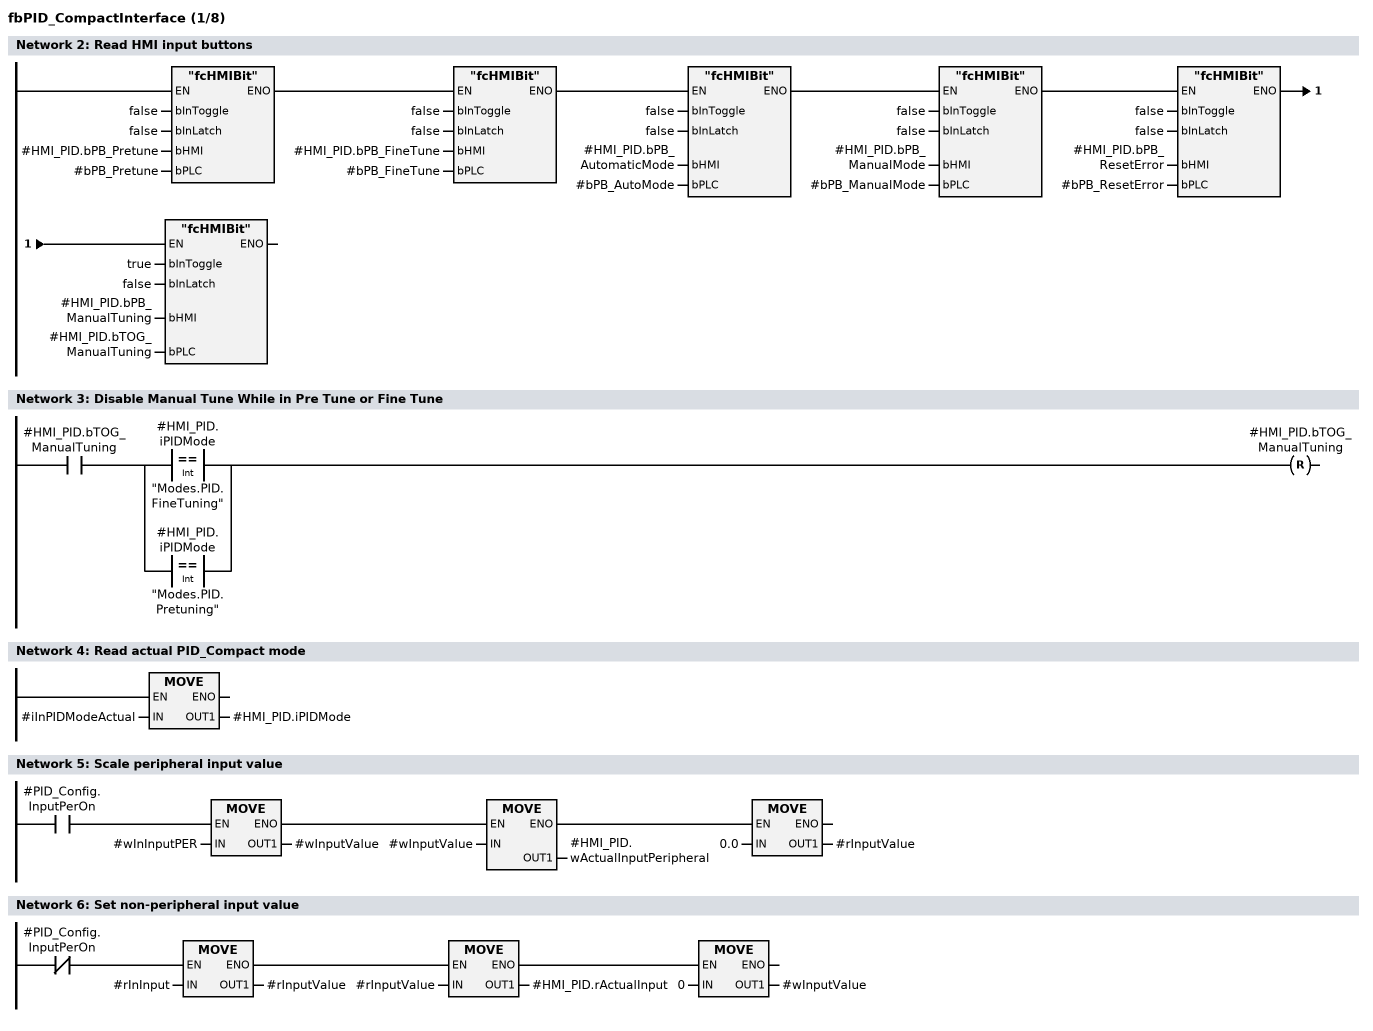
   RUNG wire#powerrail
      "fcHMIBit"(bInToggle := false, bInLatch := false, bHMI := #HMI_PID.bPB_Pretune, bPLC := #bPB_Pretune)
      "fcHMIBit"(bInToggle := false, bInLatch := false, bHMI := #HMI_PID.bPB_FineTune, bPLC := #bPB_FineTune)
      "fcHMIBit"(bInToggle := false, bInLatch := false, bHMI := #HMI_PID.bPB_AutomaticMode, bPLC := #bPB_AutoMode)
      "fcHMIBit"(bInToggle := false, bInLatch := false, bHMI := #HMI_PID.bPB_ManualMode, bPLC := #bPB_ManualMode)
      "fcHMIBit"(bInToggle := false, bInLatch := false, bHMI := #HMI_PID.bPB_ResetError, bPLC := #bPB_ResetError)
      "fcHMIBit"(bInToggle := true, bInLatch := false, bHMI := #HMI_PID.bPB_ManualTuning, bPLC := #HMI_PID.bTOG_ManualTuning)
   END_RUNG
   // the same network as SCL:
   "fcHMIBit"(bInToggle := false,
              bInLatch := false,
              bHMI := #HMI_PID.bPB_Pretune,
              bPLC := #bPB_Pretune,
              ENO => #_w1);
   "fcHMIBit"(EN := #_w1,
              bInToggle := false,
              bInLatch := false,
              bHMI := #HMI_PID.bPB_FineTune,
              bPLC := #bPB_FineTune,
              ENO => #_w2);
   "fcHMIBit"(EN := #_w2,
              bInToggle := false,
              bInLatch := false,
              bHMI := #HMI_PID.bPB_AutomaticMode,
              bPLC := #bPB_AutoMode,
              ENO => #_w3);
   "fcHMIBit"(EN := #_w3,
              bInToggle := false,
              bInLatch := false,
              bHMI := #HMI_PID.bPB_ManualMode,
              bPLC := #bPB_ManualMode,
              ENO => #_w4);
   "fcHMIBit"(EN := #_w4,
              bInToggle := false,
              bInLatch := false,
              bHMI := #HMI_PID.bPB_ResetError,
              bPLC := #bPB_ResetError,
              ENO => #_w5);
   IF #_w5 THEN
       "fcHMIBit"(bInToggle := true,
                  bInLatch := false,
                  bHMI := #HMI_PID.bPB_ManualTuning,
                  bPLC := #HMI_PID.bTOG_ManualTuning);
   END_IF;
END_REGION

REGION Network 3: Disable Manual Tune While in Pre Tune or Fine Tune
   RUNG wire#powerrail
      Contact( #HMI_PID.bTOG_ManualTuning )
      wire#w1
      { S7_Templates := "SrcType := Int" } EQ_Contact(in1 := #HMI_PID.iPIDMode, in2 := "Modes.PID.FineTuning")
      wire#w2
      R_Coil( #HMI_PID.bTOG_ManualTuning )
   END_RUNG
   RUNG wire#w1
      { S7_Templates := "SrcType := Int" } EQ_Contact(in1 := #HMI_PID.iPIDMode, in2 := "Modes.PID.Pretuning")
   END_RUNG wire#w2
   // the same network as SCL:
   IF #HMI_PID.bTOG_ManualTuning AND ((#HMI_PID.iPIDMode = "Modes.PID.FineTuning") OR (#HMI_PID.iPIDMode = "Modes.PID.Pretuning")) THEN
       #HMI_PID.bTOG_ManualTuning := FALSE;
   END_IF;
END_REGION

REGION Network 4: Read actual PID_Compact mode
   RUNG wire#powerrail
      Move(in := #iInPIDModeActual, out1 => #HMI_PID.iPIDMode)
   END_RUNG
   // the same network as SCL:
   #HMI_PID.iPIDMode := #iInPIDModeActual;
END_REGION

REGION Network 5: Scale peripheral input value
   RUNG wire#powerrail
      Contact( #PID_Config.InputPerOn )
      Move(in := #wInInputPER, out1 => #wInputValue)
      Move(in := #wInputValue, out1 => #HMI_PID.wActualInputPeripheral)
      Move(in := 0.0, out1 => #rInputValue)
   END_RUNG
   // the same network as SCL:
   IF #PID_Config.InputPerOn THEN
       #wInputValue := #wInInputPER;
       #HMI_PID.wActualInputPeripheral := #wInputValue;
       #rInputValue := 0.0;
   END_IF;
END_REGION

REGION Network 6: Set non-peripheral input value
   RUNG wire#powerrail
      I_Contact( #PID_Config.InputPerOn )
      Move(in := #rInInput, out1 => #rInputValue)
      Move(in := #rInputValue, out1 => #HMI_PID.rActualInput)
      Move(in := 0, out1 => #wInputValue)
   END_RUNG
   // the same network as SCL:
   IF NOT #PID_Config.InputPerOn THEN
       #rInputValue := #rInInput;
       #HMI_PID.rActualInput := #rInputValue;
       #wInputValue := 0;
   END_IF;
END_REGION

REGION Network 7: Check HMI tuning parameters for changes
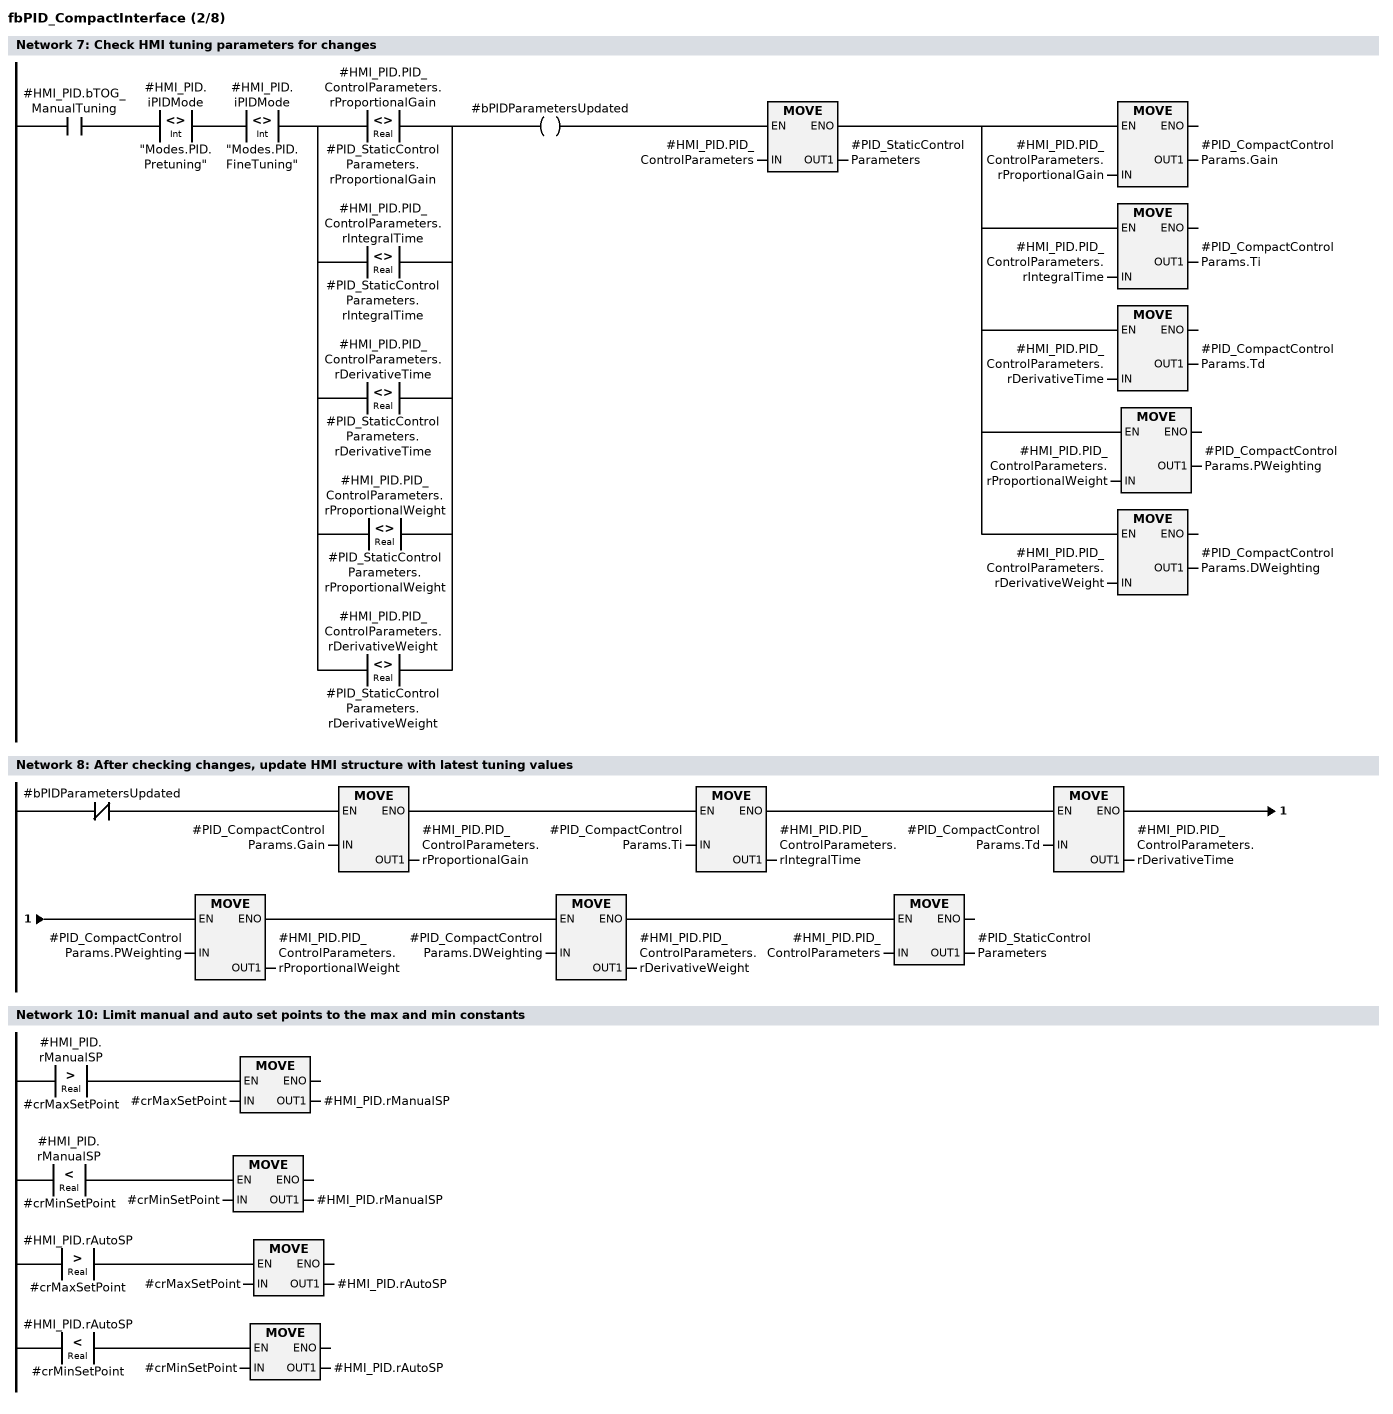
   RUNG wire#powerrail
      Contact( #HMI_PID.bTOG_ManualTuning )
      { S7_Templates := "SrcType := Int" } NE_Contact(in1 := #HMI_PID.iPIDMode, in2 := "Modes.PID.Pretuning")
      { S7_Templates := "SrcType := Int" } NE_Contact(in1 := #HMI_PID.iPIDMode, in2 := "Modes.PID.FineTuning")
      wire#w1
      { S7_Templates := "SrcType := Real" } NE_Contact(in1 := #HMI_PID.PID_ControlParameters.rProportionalGain, in2 := #PID_StaticControlParameters.rProportionalGain)
      wire#w2
      Coil( #bPIDParametersUpdated )
      Move(in := #HMI_PID.PID_ControlParameters, out1 => #PID_StaticControlParameters)
      wire#w3
      Move(in := #HMI_PID.PID_ControlParameters.rProportionalGain, out1 => #PID_CompactControlParams.Gain)
   END_RUNG
   RUNG wire#w1
      { S7_Templates := "SrcType := Real" } NE_Contact(in1 := #HMI_PID.PID_ControlParameters.rIntegralTime, in2 := #PID_StaticControlParameters.rIntegralTime)
   END_RUNG wire#w2
   RUNG wire#w1
      { S7_Templates := "SrcType := Real" } NE_Contact(in1 := #HMI_PID.PID_ControlParameters.rDerivativeTime, in2 := #PID_StaticControlParameters.rDerivativeTime)
   END_RUNG wire#w2
   RUNG wire#w1
      { S7_Templates := "SrcType := Real" } NE_Contact(in1 := #HMI_PID.PID_ControlParameters.rProportionalWeight, in2 := #PID_StaticControlParameters.rProportionalWeight)
   END_RUNG wire#w2
   RUNG wire#w1
      { S7_Templates := "SrcType := Real" } NE_Contact(in1 := #HMI_PID.PID_ControlParameters.rDerivativeWeight, in2 := #PID_StaticControlParameters.rDerivativeWeight)
   END_RUNG wire#w2
   RUNG wire#w3
      Move(in := #HMI_PID.PID_ControlParameters.rIntegralTime, out1 => #PID_CompactControlParams.Ti)
   END_RUNG
   RUNG wire#w3
      Move(in := #HMI_PID.PID_ControlParameters.rDerivativeTime, out1 => #PID_CompactControlParams.Td)
   END_RUNG
   RUNG wire#w3
      Move(in := #HMI_PID.PID_ControlParameters.rProportionalWeight, out1 => #PID_CompactControlParams.PWeighting)
   END_RUNG
   RUNG wire#w3
      Move(in := #HMI_PID.PID_ControlParameters.rDerivativeWeight, out1 => #PID_CompactControlParams.DWeighting)
   END_RUNG
   // the same network as SCL:
   #bPIDParametersUpdated := #HMI_PID.bTOG_ManualTuning AND (#HMI_PID.iPIDMode <> "Modes.PID.Pretuning") AND (#HMI_PID.iPIDMode <> "Modes.PID.FineTuning") AND ((#HMI_PID.PID_ControlParameters.rProportionalGain <> #PID_StaticControlParameters.rProportionalGain) OR (#HMI_PID.PID_ControlParameters.rIntegralTime <> #PID_StaticControlParameters.rIntegralTime) OR (#HMI_PID.PID_ControlParameters.rDerivativeTime <> #PID_StaticControlParameters.rDerivativeTime) OR (#HMI_PID.PID_ControlParameters.rProportionalWeight <> #PID_StaticControlParameters.rProportionalWeight) OR (#HMI_PID.PID_ControlParameters.rDerivativeWeight <> #PID_StaticControlParameters.rDerivativeWeight));
   IF #bPIDParametersUpdated THEN
       #PID_StaticControlParameters := #HMI_PID.PID_ControlParameters;
       #PID_CompactControlParams.Gain := #HMI_PID.PID_ControlParameters.rProportionalGain;
       #PID_CompactControlParams.Ti := #HMI_PID.PID_ControlParameters.rIntegralTime;
       #PID_CompactControlParams.Td := #HMI_PID.PID_ControlParameters.rDerivativeTime;
       #PID_CompactControlParams.PWeighting := #HMI_PID.PID_ControlParameters.rProportionalWeight;
       #PID_CompactControlParams.DWeighting := #HMI_PID.PID_ControlParameters.rDerivativeWeight;
   END_IF;
END_REGION

REGION Network 8: After checking changes, update HMI structure with latest tuning values
   RUNG wire#powerrail
      I_Contact( #bPIDParametersUpdated )
      Move(in := #PID_CompactControlParams.Gain, out1 => #HMI_PID.PID_ControlParameters.rProportionalGain)
      Move(in := #PID_CompactControlParams.Ti, out1 => #HMI_PID.PID_ControlParameters.rIntegralTime)
      Move(in := #PID_CompactControlParams.Td, out1 => #HMI_PID.PID_ControlParameters.rDerivativeTime)
      Move(in := #PID_CompactControlParams.PWeighting, out1 => #HMI_PID.PID_ControlParameters.rProportionalWeight)
      Move(in := #PID_CompactControlParams.DWeighting, out1 => #HMI_PID.PID_ControlParameters.rDerivativeWeight)
      Move(in := #HMI_PID.PID_ControlParameters, out1 => #PID_StaticControlParameters)
   END_RUNG
   // the same network as SCL:
   IF NOT #bPIDParametersUpdated THEN
       #HMI_PID.PID_ControlParameters.rProportionalGain := #PID_CompactControlParams.Gain;
       #HMI_PID.PID_ControlParameters.rIntegralTime := #PID_CompactControlParams.Ti;
       #HMI_PID.PID_ControlParameters.rDerivativeTime := #PID_CompactControlParams.Td;
       #HMI_PID.PID_ControlParameters.rProportionalWeight := #PID_CompactControlParams.PWeighting;
       #HMI_PID.PID_ControlParameters.rDerivativeWeight := #PID_CompactControlParams.DWeighting;
       #PID_StaticControlParameters := #HMI_PID.PID_ControlParameters;
   END_IF;
END_REGION

REGION Network 9: --------------------------------------------------- Control Logic ------------------------------------------------------------
END_REGION

REGION Network 10: Limit manual and auto set points to the max and min constants
   RUNG wire#powerrail
      { S7_Templates := "SrcType := Real" } GT_Contact(in1 := #HMI_PID.rManualSP, in2 := #crMaxSetPoint)
      { S7_GenerateENO := "TRUE" } Move(in := #crMaxSetPoint, out1 => #HMI_PID.rManualSP)
   END_RUNG
   RUNG wire#powerrail
      { S7_Templates := "SrcType := Real" } LT_Contact(in1 := #HMI_PID.rManualSP, in2 := #crMinSetPoint)
      { S7_GenerateENO := "TRUE" } Move(in := #crMinSetPoint, out1 => #HMI_PID.rManualSP)
   END_RUNG
   RUNG wire#powerrail
      { S7_Templates := "SrcType := Real" } GT_Contact(in1 := #HMI_PID.rAutoSP, in2 := #crMaxSetPoint)
      { S7_GenerateENO := "TRUE" } Move(in := #crMaxSetPoint, out1 => #HMI_PID.rAutoSP)
   END_RUNG
   RUNG wire#powerrail
      { S7_Templates := "SrcType := Real" } LT_Contact(in1 := #HMI_PID.rAutoSP, in2 := #crMinSetPoint)
      { S7_GenerateENO := "TRUE" } Move(in := #crMinSetPoint, out1 => #HMI_PID.rAutoSP)
   END_RUNG
   // the same network as SCL:
   IF #HMI_PID.rManualSP > #crMaxSetPoint THEN #HMI_PID.rManualSP := #crMaxSetPoint; END_IF;
   IF #HMI_PID.rManualSP < #crMinSetPoint THEN #HMI_PID.rManualSP := #crMinSetPoint; END_IF;
   IF #HMI_PID.rAutoSP > #crMaxSetPoint THEN #HMI_PID.rAutoSP := #crMaxSetPoint; END_IF;
   IF #HMI_PID.rAutoSP < #crMinSetPoint THEN #HMI_PID.rAutoSP := #crMinSetPoint; END_IF;
END_REGION

REGION Network 11: Reset errors
   // Clear all errors
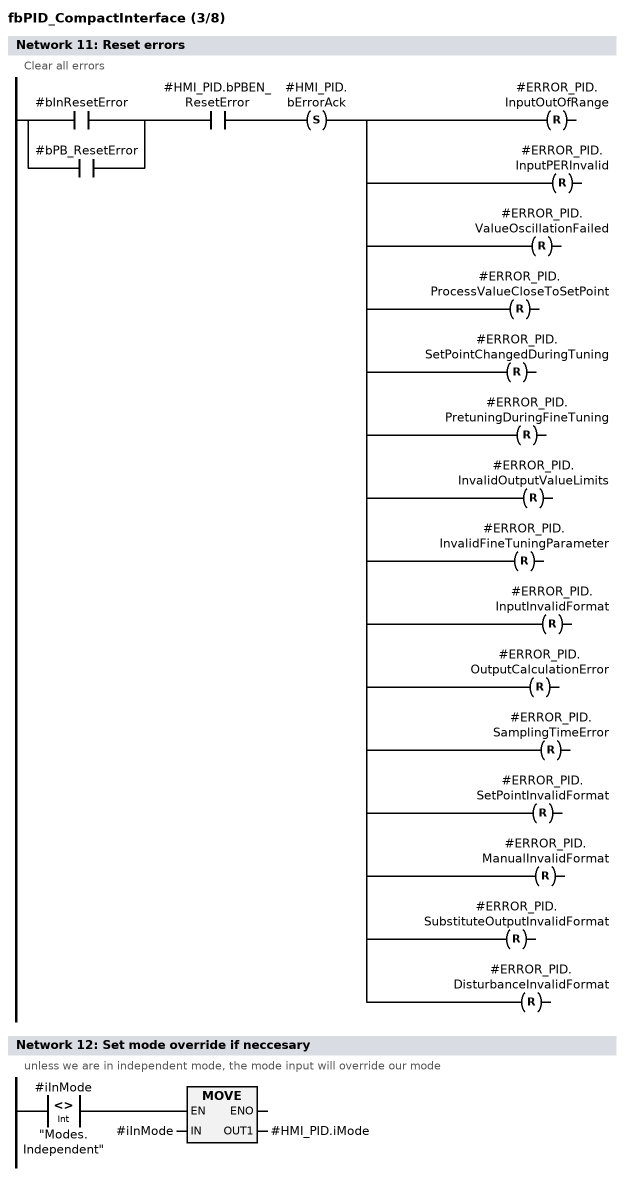
   RUNG wire#powerrail
      Contact( #bInResetError )
      wire#w1
      Contact( #HMI_PID.bPBEN_ResetError )
      S_Coil( #HMI_PID.bErrorAck )
      wire#w2
      R_Coil( #ERROR_PID.InputOutOfRange )
   END_RUNG
   RUNG wire#powerrail
      Contact( #bPB_ResetError )
   END_RUNG wire#w1
   RUNG wire#w2
      R_Coil( #ERROR_PID.InputPERInvalid )
   END_RUNG
   RUNG wire#w2
      R_Coil( #ERROR_PID.ValueOscillationFailed )
   END_RUNG
   RUNG wire#w2
      R_Coil( #ERROR_PID.ProcessValueCloseToSetPoint )
   END_RUNG
   RUNG wire#w2
      R_Coil( #ERROR_PID.SetPointChangedDuringTuning )
   END_RUNG
   RUNG wire#w2
      R_Coil( #ERROR_PID.PretuningDuringFineTuning )
   END_RUNG
   RUNG wire#w2
      R_Coil( #ERROR_PID.InvalidOutputValueLimits )
   END_RUNG
   RUNG wire#w2
      R_Coil( #ERROR_PID.InvalidFineTuningParameter )
   END_RUNG
   RUNG wire#w2
      R_Coil( #ERROR_PID.InputInvalidFormat )
   END_RUNG
   RUNG wire#w2
      R_Coil( #ERROR_PID.OutputCalculationError )
   END_RUNG
   RUNG wire#w2
      R_Coil( #ERROR_PID.SamplingTimeError )
   END_RUNG
   RUNG wire#w2
      R_Coil( #ERROR_PID.SetPointInvalidFormat )
   END_RUNG
   RUNG wire#w2
      R_Coil( #ERROR_PID.ManualInvalidFormat )
   END_RUNG
   RUNG wire#w2
      R_Coil( #ERROR_PID.SubstituteOutputInvalidFormat )
   END_RUNG
   RUNG wire#w2
      R_Coil( #ERROR_PID.DisturbanceInvalidFormat )
   END_RUNG
   // the same network as SCL:
   IF (#bInResetError OR #bPB_ResetError) AND #HMI_PID.bPBEN_ResetError THEN
       #HMI_PID.bErrorAck := TRUE;
       #ERROR_PID.InputOutOfRange := FALSE;
       #ERROR_PID.InputPERInvalid := FALSE;
       #ERROR_PID.ValueOscillationFailed := FALSE;
       #ERROR_PID.ProcessValueCloseToSetPoint := FALSE;
       #ERROR_PID.SetPointChangedDuringTuning := FALSE;
       #ERROR_PID.PretuningDuringFineTuning := FALSE;
       #ERROR_PID.InvalidOutputValueLimits := FALSE;
       #ERROR_PID.InvalidFineTuningParameter := FALSE;
       #ERROR_PID.InputInvalidFormat := FALSE;
       #ERROR_PID.OutputCalculationError := FALSE;
       #ERROR_PID.SamplingTimeError := FALSE;
       #ERROR_PID.SetPointInvalidFormat := FALSE;
       #ERROR_PID.ManualInvalidFormat := FALSE;
       #ERROR_PID.SubstituteOutputInvalidFormat := FALSE;
       #ERROR_PID.DisturbanceInvalidFormat := FALSE;
   END_IF;
END_REGION

REGION Network 12: Set mode override if neccesary
   // unless we are in independent mode, the mode input will override our mode
   RUNG wire#powerrail
      { S7_Templates := "SrcType := Int" } NE_Contact(in1 := #iInMode, in2 := "Modes.Independent")
      { S7_GenerateENO := "TRUE" } Move(in := #iInMode, out1 => #HMI_PID.iMode)
   END_RUNG
   // the same network as SCL:
   IF #iInMode <> "Modes.Independent" THEN #HMI_PID.iMode := #iInMode; END_IF;
END_REGION

REGION Network 13: Determine if auto or manual mode is active
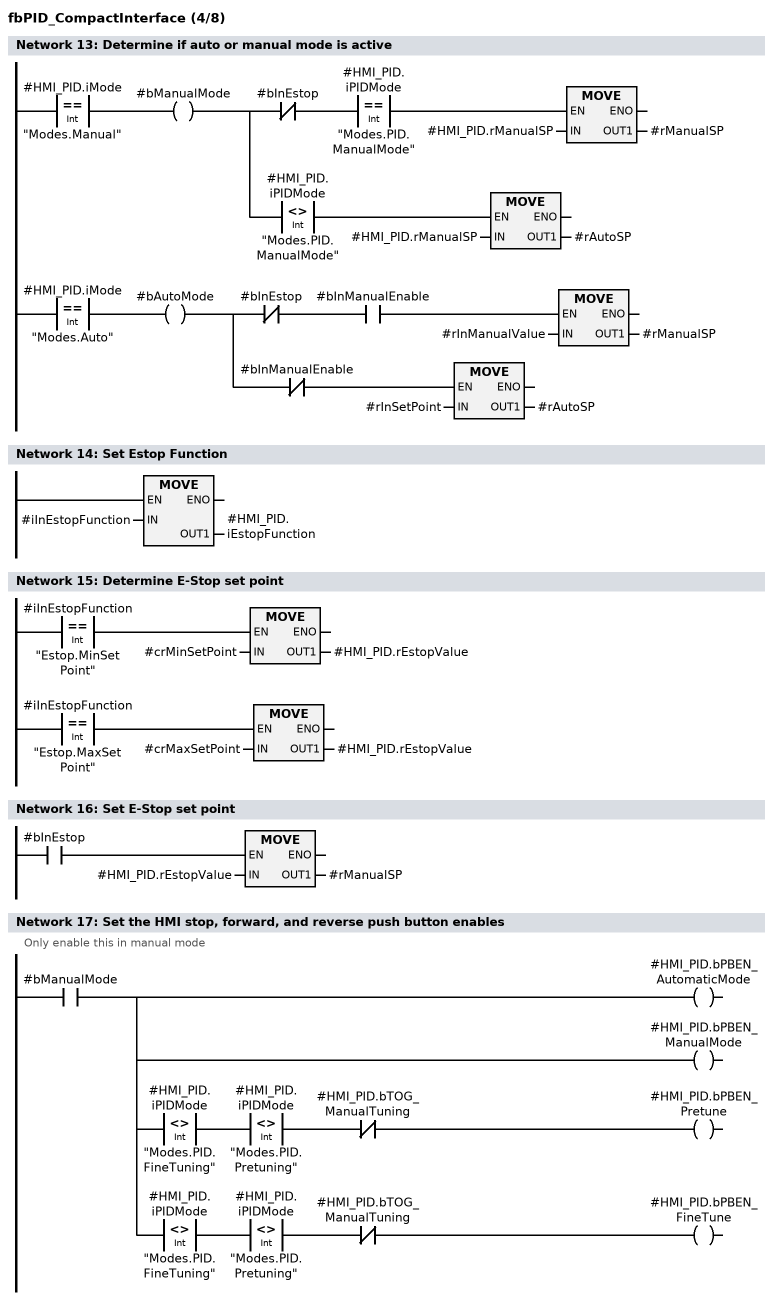
   RUNG wire#powerrail
      { S7_Templates := "SrcType := Int" } EQ_Contact(in1 := #HMI_PID.iMode, in2 := "Modes.Manual")
      Coil( #bManualMode )
      wire#w1
      I_Contact( #bInEstop )
      { S7_Templates := "SrcType := Int" } EQ_Contact(in1 := #HMI_PID.iPIDMode, in2 := "Modes.PID.ManualMode")
      { S7_GenerateENO := "TRUE" } Move(in := #HMI_PID.rManualSP, out1 => #rManualSP)
   END_RUNG
   RUNG wire#w1
      { S7_Templates := "SrcType := Int" } NE_Contact(in1 := #HMI_PID.iPIDMode, in2 := "Modes.PID.ManualMode")
      { S7_GenerateENO := "TRUE" } Move(in := #HMI_PID.rManualSP, out1 => #rAutoSP)
   END_RUNG
   RUNG wire#powerrail
      { S7_Templates := "SrcType := Int" } EQ_Contact(in1 := #HMI_PID.iMode, in2 := "Modes.Auto")
      Coil( #bAutoMode )
      wire#w2
      I_Contact( #bInEstop )
      Contact( #bInManualEnable )
      { S7_GenerateENO := "TRUE" } Move(in := #rInManualValue, out1 => #rManualSP)
   END_RUNG
   RUNG wire#w2
      I_Contact( #bInManualEnable )
      { S7_GenerateENO := "TRUE" } Move(in := #rInSetPoint, out1 => #rAutoSP)
   END_RUNG
   // the same network as SCL:
   #bManualMode := #HMI_PID.iMode = "Modes.Manual";
   IF #bManualMode AND NOT #bInEstop AND (#HMI_PID.iPIDMode = "Modes.PID.ManualMode") THEN
       #rManualSP := #HMI_PID.rManualSP;
   END_IF;
   IF #bManualMode AND (#HMI_PID.iPIDMode <> "Modes.PID.ManualMode") THEN
       #rAutoSP := #HMI_PID.rManualSP;
   END_IF;
   #bAutoMode := #HMI_PID.iMode = "Modes.Auto";
   IF #bAutoMode AND NOT #bInEstop AND #bInManualEnable THEN #rManualSP := #rInManualValue; END_IF;
   IF #bAutoMode AND NOT #bInManualEnable THEN #rAutoSP := #rInSetPoint; END_IF;
END_REGION

REGION Network 14: Set Estop Function
   RUNG wire#powerrail
      Move(in := #iInEstopFunction, out1 => #HMI_PID.iEstopFunction)
   END_RUNG
   // the same network as SCL:
   #HMI_PID.iEstopFunction := #iInEstopFunction;
END_REGION

REGION Network 15: Determine E-Stop set point
   RUNG wire#powerrail
      { S7_Templates := "SrcType := Int" } EQ_Contact(in1 := #iInEstopFunction, in2 := "Estop.MinSetPoint")
      { S7_GenerateENO := "TRUE" } Move(in := #crMinSetPoint, out1 => #HMI_PID.rEstopValue)
   END_RUNG
   RUNG wire#powerrail
      { S7_Templates := "SrcType := Int" } EQ_Contact(in1 := #iInEstopFunction, in2 := "Estop.MaxSetPoint")
      { S7_GenerateENO := "TRUE" } Move(in := #crMaxSetPoint, out1 => #HMI_PID.rEstopValue)
   END_RUNG
   // the same network as SCL:
   IF #iInEstopFunction = "Estop.MinSetPoint" THEN #HMI_PID.rEstopValue := #crMinSetPoint; END_IF;
   IF #iInEstopFunction = "Estop.MaxSetPoint" THEN #HMI_PID.rEstopValue := #crMaxSetPoint; END_IF;
END_REGION

REGION Network 16: Set E-Stop set point
   RUNG wire#powerrail
      Contact( #bInEstop )
      { S7_GenerateENO := "TRUE" } Move(in := #HMI_PID.rEstopValue, out1 => #rManualSP)
   END_RUNG
   // the same network as SCL:
   IF #bInEstop THEN #rManualSP := #HMI_PID.rEstopValue; END_IF;
END_REGION

REGION Network 17: Set the HMI stop, forward, and reverse push button enables
   // Only enable this in manual mode
   RUNG wire#powerrail
      Contact( #bManualMode )
      wire#w1
      Coil( #HMI_PID.bPBEN_AutomaticMode )
   END_RUNG
   RUNG wire#w1
      Coil( #HMI_PID.bPBEN_ManualMode )
   END_RUNG
   RUNG wire#w1
      { S7_Templates := "SrcType := Int" } NE_Contact(in1 := #HMI_PID.iPIDMode, in2 := "Modes.PID.FineTuning")
      { S7_Templates := "SrcType := Int" } NE_Contact(in1 := #HMI_PID.iPIDMode, in2 := "Modes.PID.Pretuning")
      I_Contact( #HMI_PID.bTOG_ManualTuning )
      Coil( #HMI_PID.bPBEN_Pretune )
   END_RUNG
   RUNG wire#w1
      { S7_Templates := "SrcType := Int" } NE_Contact(in1 := #HMI_PID.iPIDMode, in2 := "Modes.PID.FineTuning")
      { S7_Templates := "SrcType := Int" } NE_Contact(in1 := #HMI_PID.iPIDMode, in2 := "Modes.PID.Pretuning")
      I_Contact( #HMI_PID.bTOG_ManualTuning )
      Coil( #HMI_PID.bPBEN_FineTune )
   END_RUNG
   // the same network as SCL:
   #HMI_PID.bPBEN_AutomaticMode := #bManualMode;
   #HMI_PID.bPBEN_ManualMode := #bManualMode;
   #HMI_PID.bPBEN_Pretune := #bManualMode AND (#HMI_PID.iPIDMode <> "Modes.PID.FineTuning") AND (#HMI_PID.iPIDMode <> "Modes.PID.Pretuning") AND NOT #HMI_PID.bTOG_ManualTuning;
   #HMI_PID.bPBEN_FineTune := #bManualMode AND (#HMI_PID.iPIDMode <> "Modes.PID.FineTuning") AND (#HMI_PID.iPIDMode <> "Modes.PID.Pretuning") AND NOT #HMI_PID.bTOG_ManualTuning;
END_REGION

REGION Network 18: Enable the reset error pushbutton if there is an error
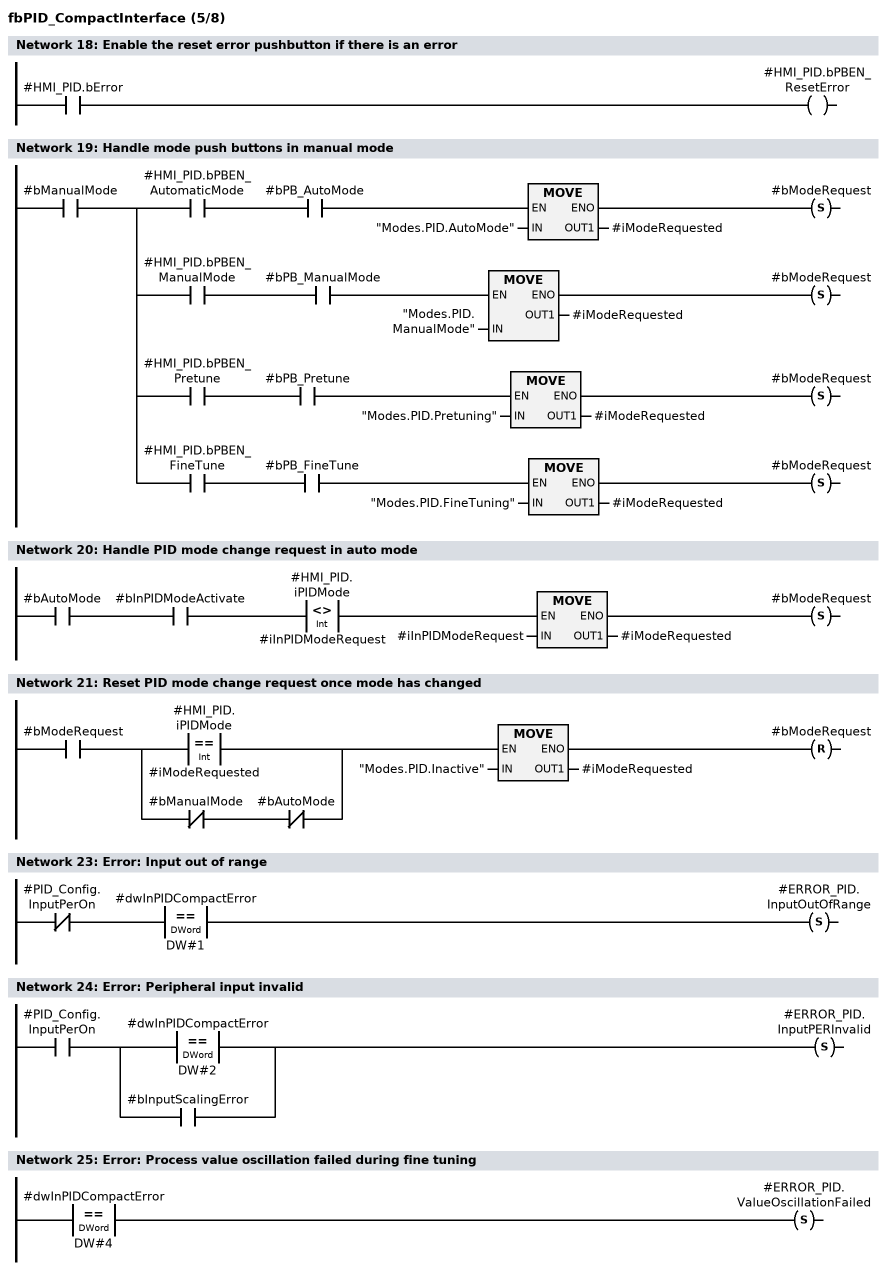
   RUNG wire#powerrail
      Contact( #HMI_PID.bError )
      Coil( #HMI_PID.bPBEN_ResetError )
   END_RUNG
   // the same network as SCL:
   #HMI_PID.bPBEN_ResetError := #HMI_PID.bError;
END_REGION

REGION Network 19: Handle mode push buttons in manual mode
   RUNG wire#powerrail
      Contact( #bManualMode )
      wire#w1
      Contact( #HMI_PID.bPBEN_AutomaticMode )
      Contact( #bPB_AutoMode )
      Move(in := "Modes.PID.AutoMode", out1 => #iModeRequested)
      S_Coil( #bModeRequest )
   END_RUNG
   RUNG wire#w1
      Contact( #HMI_PID.bPBEN_ManualMode )
      Contact( #bPB_ManualMode )
      Move(in := "Modes.PID.ManualMode", out1 => #iModeRequested)
      S_Coil( #bModeRequest )
   END_RUNG
   RUNG wire#w1
      Contact( #HMI_PID.bPBEN_Pretune )
      Contact( #bPB_Pretune )
      Move(in := "Modes.PID.Pretuning", out1 => #iModeRequested)
      S_Coil( #bModeRequest )
   END_RUNG
   RUNG wire#w1
      Contact( #HMI_PID.bPBEN_FineTune )
      Contact( #bPB_FineTune )
      Move(in := "Modes.PID.FineTuning", out1 => #iModeRequested)
      S_Coil( #bModeRequest )
   END_RUNG
   // the same network as SCL:
   IF #bManualMode AND #HMI_PID.bPBEN_AutomaticMode AND #bPB_AutoMode THEN
       #iModeRequested := "Modes.PID.AutoMode";
       #bModeRequest := TRUE;
   END_IF;
   IF #bManualMode AND #HMI_PID.bPBEN_ManualMode AND #bPB_ManualMode THEN
       #iModeRequested := "Modes.PID.ManualMode";
       #bModeRequest := TRUE;
   END_IF;
   IF #bManualMode AND #HMI_PID.bPBEN_Pretune AND #bPB_Pretune THEN
       #iModeRequested := "Modes.PID.Pretuning";
       #bModeRequest := TRUE;
   END_IF;
   IF #bManualMode AND #HMI_PID.bPBEN_FineTune AND #bPB_FineTune THEN
       #iModeRequested := "Modes.PID.FineTuning";
       #bModeRequest := TRUE;
   END_IF;
END_REGION

REGION Network 20: Handle PID mode change request in auto mode
   RUNG wire#powerrail
      Contact( #bAutoMode )
      Contact( #bInPIDModeActivate )
      { S7_Templates := "SrcType := Int" } NE_Contact(in1 := #HMI_PID.iPIDMode, in2 := #iInPIDModeRequest)
      Move(in := #iInPIDModeRequest, out1 => #iModeRequested)
      S_Coil( #bModeRequest )
   END_RUNG
   // the same network as SCL:
   IF #bAutoMode AND #bInPIDModeActivate AND (#HMI_PID.iPIDMode <> #iInPIDModeRequest) THEN
       #iModeRequested := #iInPIDModeRequest;
       #bModeRequest := TRUE;
   END_IF;
END_REGION

REGION Network 21: Reset PID mode change request once mode has changed
   RUNG wire#powerrail
      Contact( #bModeRequest )
      wire#w1
      { S7_Templates := "SrcType := Int" } EQ_Contact(in1 := #HMI_PID.iPIDMode, in2 := #iModeRequested)
      wire#w2
      Move(in := "Modes.PID.Inactive", out1 => #iModeRequested)
      R_Coil( #bModeRequest )
   END_RUNG
   RUNG wire#w1
      I_Contact( #bManualMode )
      I_Contact( #bAutoMode )
   END_RUNG wire#w2
   // the same network as SCL:
   #_w1 := #bModeRequest AND ((#HMI_PID.iPIDMode = #iModeRequested) OR (NOT #bManualMode AND NOT #bAutoMode));
   IF #_w1 THEN
       #iModeRequested := "Modes.PID.Inactive";
       #bModeRequest := FALSE;
   END_IF;
END_REGION

REGION Network 22: --------------------------------------------------------- Errors ------------------------------------------------------------------
END_REGION

REGION Network 23: Error: Input out of range
   RUNG wire#powerrail
      I_Contact( #PID_Config.InputPerOn )
      { S7_Templates := "SrcType := DWord" } EQ_Contact(in1 := #dwInPIDCompactError, in2 := DW#1)
      S_Coil( #ERROR_PID.InputOutOfRange )
   END_RUNG
   // the same network as SCL:
   IF NOT #PID_Config.InputPerOn AND (#dwInPIDCompactError = DW#1) THEN
       #ERROR_PID.InputOutOfRange := TRUE;
   END_IF;
END_REGION

REGION Network 24: Error: Peripheral input invalid
   RUNG wire#powerrail
      Contact( #PID_Config.InputPerOn )
      wire#w1
      { S7_Templates := "SrcType := DWord" } EQ_Contact(in1 := #dwInPIDCompactError, in2 := DW#2)
      wire#w2
      S_Coil( #ERROR_PID.InputPERInvalid )
   END_RUNG
   RUNG wire#w1
      Contact( #bInputScalingError )
   END_RUNG wire#w2
   // the same network as SCL:
   IF #PID_Config.InputPerOn AND ((#dwInPIDCompactError = DW#2) OR #bInputScalingError) THEN
       #ERROR_PID.InputPERInvalid := TRUE;
   END_IF;
END_REGION

REGION Network 25: Error: Process value oscillation failed during fine tuning
   RUNG wire#powerrail
      { S7_Templates := "SrcType := DWord" } EQ_Contact(in1 := #dwInPIDCompactError, in2 := DW#4)
      S_Coil( #ERROR_PID.ValueOscillationFailed )
   END_RUNG
   // the same network as SCL:
   IF #dwInPIDCompactError = DW#4 THEN #ERROR_PID.ValueOscillationFailed := TRUE; END_IF;
END_REGION

REGION Network 26: Error: Process value too close to set point for pretuning
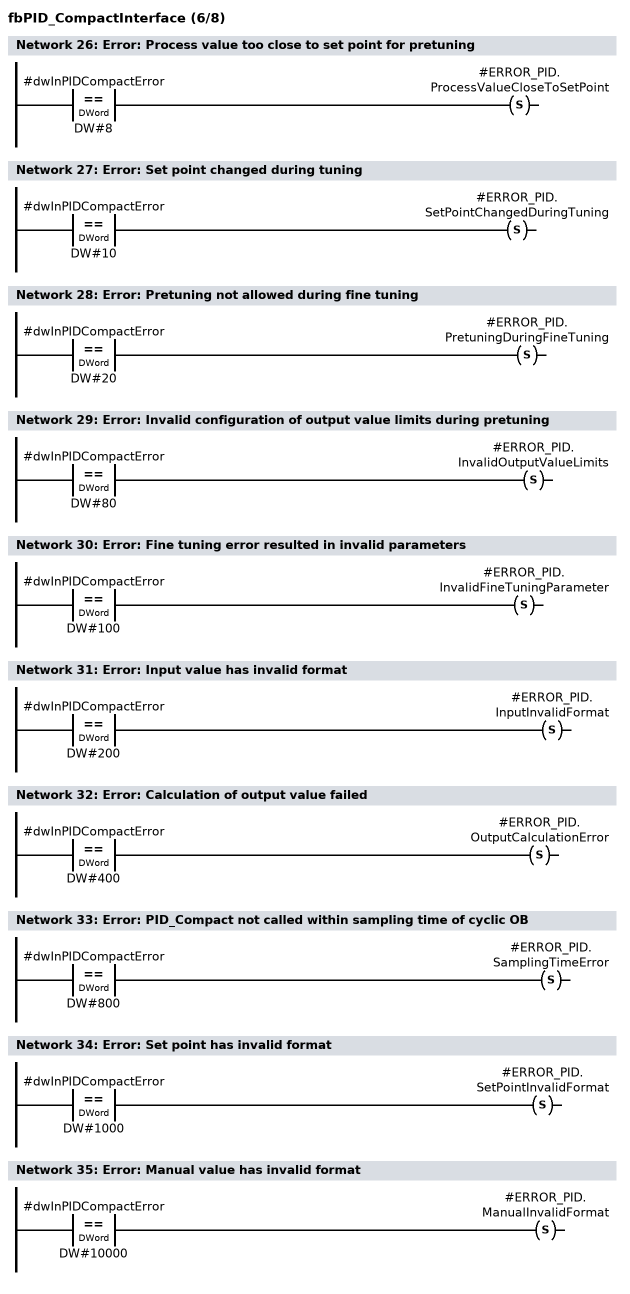
   RUNG wire#powerrail
      { S7_Templates := "SrcType := DWord" } EQ_Contact(in1 := #dwInPIDCompactError, in2 := DW#8)
      S_Coil( #ERROR_PID.ProcessValueCloseToSetPoint )
   END_RUNG
   // the same network as SCL:
   IF #dwInPIDCompactError = DW#8 THEN #ERROR_PID.ProcessValueCloseToSetPoint := TRUE; END_IF;
END_REGION

REGION Network 27: Error: Set point changed during tuning
   RUNG wire#powerrail
      { S7_Templates := "SrcType := DWord" } EQ_Contact(in1 := #dwInPIDCompactError, in2 := DW#10)
      S_Coil( #ERROR_PID.SetPointChangedDuringTuning )
   END_RUNG
   // the same network as SCL:
   IF #dwInPIDCompactError = DW#10 THEN #ERROR_PID.SetPointChangedDuringTuning := TRUE; END_IF;
END_REGION

REGION Network 28: Error: Pretuning not allowed during fine tuning
   RUNG wire#powerrail
      { S7_Templates := "SrcType := DWord" } EQ_Contact(in1 := #dwInPIDCompactError, in2 := DW#20)
      S_Coil( #ERROR_PID.PretuningDuringFineTuning )
   END_RUNG
   // the same network as SCL:
   IF #dwInPIDCompactError = DW#20 THEN #ERROR_PID.PretuningDuringFineTuning := TRUE; END_IF;
END_REGION

REGION Network 29: Error: Invalid configuration of output value limits during pretuning
   RUNG wire#powerrail
      { S7_Templates := "SrcType := DWord" } EQ_Contact(in1 := #dwInPIDCompactError, in2 := DW#80)
      S_Coil( #ERROR_PID.InvalidOutputValueLimits )
   END_RUNG
   // the same network as SCL:
   IF #dwInPIDCompactError = DW#80 THEN #ERROR_PID.InvalidOutputValueLimits := TRUE; END_IF;
END_REGION

REGION Network 30: Error: Fine tuning error resulted in invalid parameters
   RUNG wire#powerrail
      { S7_Templates := "SrcType := DWord" } EQ_Contact(in1 := #dwInPIDCompactError, in2 := DW#100)
      S_Coil( #ERROR_PID.InvalidFineTuningParameter )
   END_RUNG
   // the same network as SCL:
   IF #dwInPIDCompactError = DW#100 THEN #ERROR_PID.InvalidFineTuningParameter := TRUE; END_IF;
END_REGION

REGION Network 31: Error: Input value has invalid format
   RUNG wire#powerrail
      { S7_Templates := "SrcType := DWord" } EQ_Contact(in1 := #dwInPIDCompactError, in2 := DW#200)
      S_Coil( #ERROR_PID.InputInvalidFormat )
   END_RUNG
   // the same network as SCL:
   IF #dwInPIDCompactError = DW#200 THEN #ERROR_PID.InputInvalidFormat := TRUE; END_IF;
END_REGION

REGION Network 32: Error: Calculation of output value failed
   RUNG wire#powerrail
      { S7_Templates := "SrcType := DWord" } EQ_Contact(in1 := #dwInPIDCompactError, in2 := DW#400)
      S_Coil( #ERROR_PID.OutputCalculationError )
   END_RUNG
   // the same network as SCL:
   IF #dwInPIDCompactError = DW#400 THEN #ERROR_PID.OutputCalculationError := TRUE; END_IF;
END_REGION

REGION Network 33: Error: PID_Compact not called within sampling time of cyclic OB
   RUNG wire#powerrail
      { S7_Templates := "SrcType := DWord" } EQ_Contact(in1 := #dwInPIDCompactError, in2 := DW#800)
      S_Coil( #ERROR_PID.SamplingTimeError )
   END_RUNG
   // the same network as SCL:
   IF #dwInPIDCompactError = DW#800 THEN #ERROR_PID.SamplingTimeError := TRUE; END_IF;
END_REGION

REGION Network 34: Error: Set point has invalid format
   RUNG wire#powerrail
      { S7_Templates := "SrcType := DWord" } EQ_Contact(in1 := #dwInPIDCompactError, in2 := DW#1000)
      S_Coil( #ERROR_PID.SetPointInvalidFormat )
   END_RUNG
   // the same network as SCL:
   IF #dwInPIDCompactError = DW#1000 THEN #ERROR_PID.SetPointInvalidFormat := TRUE; END_IF;
END_REGION

REGION Network 35: Error: Manual value has invalid format
   RUNG wire#powerrail
      { S7_Templates := "SrcType := DWord" } EQ_Contact(in1 := #dwInPIDCompactError, in2 := DW#10000)
      S_Coil( #ERROR_PID.ManualInvalidFormat )
   END_RUNG
   // the same network as SCL:
   IF #dwInPIDCompactError = DW#10000 THEN #ERROR_PID.ManualInvalidFormat := TRUE; END_IF;
END_REGION

REGION Network 36: Error: Substitute Output has invalid format